   "Cooling System Operating" : Bool = PLC "68_Sys_Status_Data".CSW_IL_PRES_IN_RNG AT %DB1.DBX0.0, 1 s
   "Correct Phase Rotation" : Bool = PLC "10_DI_Data".MCCP_5PG1_OK AT %DB1.DBX0.0, 1 s
   "CSW Drain Valve Closed" : Bool = PLC "10_DI_Data".CV322_CLSD AT %DB1.DBX0.0, 1 s
   "CSW Drain Valve Control" : Bool = PLC "14_DQ_Data".CV321_322_CNTRL AT %DB1.DBX0.0, 1 s
   "CSW Drain Valve Open" : Bool = PLC "10_DI_Data".CV322_OPN AT %DB1.DBX0.0, 1 s
   "CSW Pump Control" : Bool = PLC "51_SLAVE_STATUS".P301_ENBLD AT %DB51.DBX14.3, 1 s
   "CSW Pump Enabled" : Bool = PLC "10 DI_DATA".P301_ENBLD AT %DB1.DBX0.0, 1 s
   "CSW Pump Tripped" : Bool = PLC "10 DI_DATA".P301_TRIPPED AT %DB1.DBX0.0, 1 s
   "CSW Valve Closed" : Bool = PLC "10_DI_Data".CV311_CLSD AT %DB1.DBW0, 1 s
   "CSW Valve Control" : Bool = PLC "14_DQ_Data".CV311_312_CNTRL AT %DB1.DBX0.0, 1 s
   "CSW Valve Open" : Bool = PLC "10_DI_Data".CV311_OPN AT %DB1.DBW0, 1 s
   "Current User" : WString[15] AT %DB1.DBX0.0
   "CV312 Present" : Bool = PLC "80_From_HMI".CV312_PRSNT AT %DB1.DBX0.0, 1 s
   "CV401 - IG Supply Valve Closed" : Bool = PLC "10_DI_Data".CV401_CLSD AT %DB1.DBX0.0, 1 s
   "CV401 - IG Supply Valve Control" : Bool = PLC "14_DQ_Data".CV401_CNTRL AT %DB1.DBX0.0, 1 s
   "CV401 - IG Supply Valve Opened" : Bool = PLC "10_DI_Data".CV401_OPN AT %DB1.DBX0.0, 1 s
   "CV403 - IG Vent Valve Position Feedback Scaled" : Real = PLC "12_AI_Data".CV403_SCALED AT %DB1.DBX0.0, 1 s
   "CV431 Present" : Bool = PLC "80_From_HMI".CV431_PRSNT AT %DB1.DBX0.0, 1 s
   "CV431/432 CB/BWTS Valve" : Bool = PLC "14_DQ_Data".CV431_432_CNTRL AT %DB1.DBX0.0, 1 s
   "CV432 Present" : Bool = PLC "80_From_HMI".CV432_PRSNT AT %DB1.DBX0.0, 1 s
   "Data To IGG PLC_Data_Fuel Oil System Proved" : Bool = PLC "68_Sys_Status_Data".FUEL_PRES_IN_RNG AT %DB1.DBX0.0, 1 s
   "Data To IGG PLC_Data_VSD Fault Flag" : Bool = PLC "10_DI_Data".E139_VSD_FLT AT %DB1.DBX0.0, 1 s
   "Data_From BC PLC_Data_IA Compressor Running" : Bool = PLC "68_Sys_Status_Data".IA_PRES_IN_RNG AT %DB1.DBX0.0, 1 s
   "Data_To_BC PLC_Data_Cooling Water System Proved" : Bool = PLC "10_DI_Data".CV311_OPN AT %DB1.DBX0.0, 1 s
   "db_time_sync_time_local_READ" : LDT = PLC db_time_sync_time_local_READ AT %M4.0, 1 s
   "db_time_sync_time_system_READ" : LDT = PLC db_time_sync_time_system_READ AT %M2.0, 1 s
   "DTB Valve Closed" : Bool = PLC "10_DI_Data".CV321_CLSD AT %DB1.DBX0.0, 1 s
   "DTB Valve Opened" : Bool = PLC "10_DI_Data".CV321_OPN AT %DB1.DBX0.0, 1 s
   "Evolving Setpoint_DB_LevelBetter" : Bool = PLC "Evolving Setpoint_DB".LevelBetter, 1 s
   "External Shutdown" : Bool = PLC "10 DI_DATA".ESD_OK AT %DB1.DBX0.0, 1 s
   "FDU Power Healthy" : Bool = PLC "10 DI_DATA".FD001_PWR_OK AT %DB1.DBX0.0, 1 s
   "FIT417_1S__ALM_ANALOG_DB_HIGH LEVEL VALUE (H)" : Real = PLC "FIT417_1S__ALM_ANALOG_DB"."HIGH LEVEL VALUE (H)" AT %DB2090.DBD30, 1 s
   "FIT417_1S__ALM_ANALOG_DB_LOW LEVEL VALUE (L)" : Real = PLC "FIT417_1S__ALM_ANALOG_DB"."LOW LEVEL VALUE (L)" AT %DB2090.DBD26, 1 s
   "FIT417_1S__ALM_ANALOG_DB_VERY HIGH LEVEL VALUE (HH)" : Real = PLC "FIT417_1S__ALM_ANALOG_DB"."VERY HIGH LEVEL VALUE (HH)" AT %DB2090.DBD34, 1 s
   "FIT417_1S__ALM_ANALOG_DB_VERY LOW LEVEL VALUE (LL)" : Real = PLC "FIT417_1S__ALM_ANALOG_DB"."VERY LOW LEVEL VALUE (LL)" AT %DB2090.DBD22, 1 s
   "FIT417_2S_ALM_ANALOG_DB_HIGH LEVEL VALUE (H)" : Real = PLC FIT417_2S_ALM_ANALOG_DB."HIGH LEVEL VALUE (H)" AT %DB2066.DBD30, 1 s
   "FIT417_2S_ALM_ANALOG_DB_LOW LEVEL VALUE (L)" : Real = PLC FIT417_2S_ALM_ANALOG_DB."LOW LEVEL VALUE (L)" AT %DB2066.DBD26, 1 s
   "FIT417_2S_ALM_ANALOG_DB_VERY HIGH LEVEL VALUE (HH)" : Real = PLC FIT417_2S_ALM_ANALOG_DB."VERY HIGH LEVEL VALUE (HH)" AT %DB2066.DBD34, 1 s
   "FIT417_2S_ALM_ANALOG_DB_VERY LOW LEVEL VALUE (LL)" : Real = PLC FIT417_2S_ALM_ANALOG_DB."VERY LOW LEVEL VALUE (LL)" AT %DB2066.DBD22, 1 s
   "FIT417_3S_ALM_ANALOG_DB_HIGH LEVEL VALUE (H)" : Real = PLC FIT417_3S_ALM_ANALOG_DB."HIGH LEVEL VALUE (H)" AT %DB2092.DBD30, 1 s
   "FIT417_3S_ALM_ANALOG_DB_LOW LEVEL VALUE (L)" : Real = PLC FIT417_3S_ALM_ANALOG_DB."LOW LEVEL VALUE (L)" AT %DB2092.DBD26, 1 s
   "FIT417_3S_ALM_ANALOG_DB_VERY HIGH LEVEL VALUE (HH)" : Real = PLC FIT417_3S_ALM_ANALOG_DB."VERY HIGH LEVEL VALUE (HH)" AT %DB2092.DBD34, 1 s
   "FIT417_3S_ALM_ANALOG_DB_VERY LOW LEVEL VALUE (LL)" : Real = PLC FIT417_3S_ALM_ANALOG_DB."VERY LOW LEVEL VALUE (LL)" AT %DB2092.DBD22, 1 s
   "FIT417_4S_ALM_ANALOG_DB_HIGH LEVEL VALUE (H)" : Real = PLC FIT417_4S_ALM_ANALOG_DB."HIGH LEVEL VALUE (H)" AT %DB2094.DBD30, 1 s
   "FIT417_4S_ALM_ANALOG_DB_LOW LEVEL VALUE (L)" : Real = PLC FIT417_4S_ALM_ANALOG_DB."LOW LEVEL VALUE (L)" AT %DB2094.DBD26, 1 s
   "FIT417_4S_ALM_ANALOG_DB_VERY HIGH LEVEL VALUE (HH)" : Real = PLC FIT417_4S_ALM_ANALOG_DB."VERY HIGH LEVEL VALUE (HH)" AT %DB2094.DBD34, 1 s
   "FIT417_4S_ALM_ANALOG_DB_VERY LOW LEVEL VALUE (LL)" : Real = PLC FIT417_4S_ALM_ANALOG_DB."VERY LOW LEVEL VALUE (LL)" AT %DB2094.DBD22, 1 s
   "FIT417_5S_ALM_ANALOG_DB_HIGH LEVEL VALUE (H)" : Real = PLC FIT417_5S_ALM_ANALOG_DB."HIGH LEVEL VALUE (H)" AT %DB2096.DBD30, 1 s
   "FIT417_5S_ALM_ANALOG_DB_LOW LEVEL VALUE (L)" : Real = PLC FIT417_5S_ALM_ANALOG_DB."LOW LEVEL VALUE (L)" AT %DB2096.DBD26, 1 s
   "FIT417_5S_ALM_ANALOG_DB_VERY HIGH LEVEL VALUE (HH)" : Real = PLC FIT417_5S_ALM_ANALOG_DB."VERY HIGH LEVEL VALUE (HH)" AT %DB2096.DBD34, 1 s
   "FIT417_5S_ALM_ANALOG_DB_VERY LOW LEVEL VALUE (LL)" : Real = PLC FIT417_5S_ALM_ANALOG_DB."VERY LOW LEVEL VALUE (LL)" AT %DB2096.DBD22, 1 s
   "FIT417_6S_ALM_ANALOG_DB_HIGH LEVEL VALUE (H)" : Real = PLC FIT417_6S_ALM_ANALOG_DB."HIGH LEVEL VALUE (H)" AT %DB2098.DBD30, 1 s
   "FIT417_6S_ALM_ANALOG_DB_LOW LEVEL VALUE (L)" : Real = PLC FIT417_6S_ALM_ANALOG_DB."LOW LEVEL VALUE (L)" AT %DB2098.DBD26, 1 s
   "FIT417_6S_ALM_ANALOG_DB_VERY HIGH LEVEL VALUE (HH)" : Real = PLC FIT417_6S_ALM_ANALOG_DB."VERY HIGH LEVEL VALUE (HH)" AT %DB2098.DBD34, 1 s
   "FIT417_6S_ALM_ANALOG_DB_VERY LOW LEVEL VALUE (LL)" : Real = PLC FIT417_6S_ALM_ANALOG_DB."VERY LOW LEVEL VALUE (LL)" AT %DB2098.DBD22, 1 s
   "FIT417_APT_ALM_ANALOG_DB_HIGH LEVEL VALUE (H)" : Real = PLC FIT417_APT_ALM_ANALOG_DB."HIGH LEVEL VALUE (H)" AT %DB2099.DBD30, 1 s
   "FIT417_APT_ALM_ANALOG_DB_LOW LEVEL VALUE (L)" : Real = PLC FIT417_APT_ALM_ANALOG_DB."LOW LEVEL VALUE (L)" AT %DB2099.DBD26, 1 s
   "FIT417_APT_ALM_ANALOG_DB_VERY HIGH LEVEL VALUE (HH)" : Real = PLC FIT417_APT_ALM_ANALOG_DB."VERY HIGH LEVEL VALUE (HH)" AT %DB2099.DBD34, 1 s
   "FIT417_APT_ALM_ANALOG_DB_VERY LOW LEVEL VALUE (LL)" : Real = PLC FIT417_APT_ALM_ANALOG_DB."VERY LOW LEVEL VALUE (LL)" AT %DB2099.DBD22, 1 s
   "FIT418_1P__ALM_ANALOG_DB_HIGH LEVEL VALUE (H)" : Real = PLC "FIT418_1P__ALM_ANALOG_DB"."HIGH LEVEL VALUE (H)" AT %DB2089.DBD30, 1 s
   "FIT418_1P__ALM_ANALOG_DB_LOW LEVEL VALUE (L)" : Real = PLC "FIT418_1P__ALM_ANALOG_DB"."LOW LEVEL VALUE (L)" AT %DB2089.DBD26, 1 s
   "FIT418_1P__ALM_ANALOG_DB_VERY HIGH LEVEL VALUE (HH)" : Real = PLC "FIT418_1P__ALM_ANALOG_DB"."VERY HIGH LEVEL VALUE (HH)" AT %DB2089.DBD34, 1 s
   "FIT418_1P__ALM_ANALOG_DB_VERY LOW LEVEL VALUE (LL)" : Real = PLC "FIT418_1P__ALM_ANALOG_DB"."VERY LOW LEVEL VALUE (LL)" AT %DB2089.DBD22, 1 s
   "FIT418_2P_ALM_ANALOG_DB_ALARM L" : Bool = PLC FIT418_2P_ALM_ANALOG_DB."ALARM L" AT %DB2064.DBX48.2, 1 s
   "FIT418_2P_ALM_ANALOG_DB_HIGH LEVEL VALUE (H)" : Real = PLC FIT418_2P_ALM_ANALOG_DB."HIGH LEVEL VALUE (H)" AT %DB2064.DBD30, 1 s
   "FIT418_2P_ALM_ANALOG_DB_LOW LEVEL VALUE (L)" : Real = PLC FIT418_2P_ALM_ANALOG_DB."LOW LEVEL VALUE (L)" AT %DB2064.DBD26, 1 s
   "FIT418_2P_ALM_ANALOG_DB_VERY HIGH LEVEL VALUE (HH)" : Real = PLC FIT418_2P_ALM_ANALOG_DB."VERY HIGH LEVEL VALUE (HH)" AT %DB2064.DBD34, 1 s
   "FIT418_2P_ALM_ANALOG_DB_VERY LOW LEVEL VALUE (LL)" : Real = PLC FIT418_2P_ALM_ANALOG_DB."VERY LOW LEVEL VALUE (LL)" AT %DB2064.DBD22, 1 s
   "FIT418_3P__ALM_ANALOG_DB_HIGH LEVEL VALUE (H)" : Real = PLC "FIT418_3P__ALM_ANALOG_DB"."HIGH LEVEL VALUE (H)" AT %DB2091.DBD30, 1 s
   "FIT418_3P__ALM_ANALOG_DB_LOW LEVEL VALUE (L)" : Real = PLC "FIT418_3P__ALM_ANALOG_DB"."LOW LEVEL VALUE (L)" AT %DB2091.DBD26, 1 s
   "FIT418_3P__ALM_ANALOG_DB_VERY HIGH LEVEL VALUE (HH)" : Real = PLC "FIT418_3P__ALM_ANALOG_DB"."VERY HIGH LEVEL VALUE (HH)" AT %DB2091.DBD34, 1 s
   "FIT418_3P__ALM_ANALOG_DB_VERY LOW LEVEL VALUE (LL)" : Real = PLC "FIT418_3P__ALM_ANALOG_DB"."VERY LOW LEVEL VALUE (LL)" AT %DB2091.DBD22, 1 s
   "FIT418_4P__ALM_ANALOG_DB_HIGH LEVEL VALUE (H)" : Real = PLC "FIT418_4P__ALM_ANALOG_DB"."HIGH LEVEL VALUE (H)" AT %DB2093.DBD30, 1 s
   "FIT418_4P__ALM_ANALOG_DB_LOW LEVEL VALUE (L)" : Real = PLC "FIT418_4P__ALM_ANALOG_DB"."LOW LEVEL VALUE (L)" AT %DB2093.DBD26, 1 s
   "FIT418_4P__ALM_ANALOG_DB_VERY HIGH LEVEL VALUE (HH)" : Real = PLC "FIT418_4P__ALM_ANALOG_DB"."VERY HIGH LEVEL VALUE (HH)" AT %DB2093.DBD34, 1 s
   "FIT418_4P__ALM_ANALOG_DB_VERY LOW LEVEL VALUE (LL)" : Real = PLC "FIT418_4P__ALM_ANALOG_DB"."VERY LOW LEVEL VALUE (LL)" AT %DB2093.DBD22, 1 s
   "FIT418_5P__ALM_ANALOG_DB_HIGH LEVEL VALUE (H)" : Real = PLC "FIT418_5P__ALM_ANALOG_DB"."HIGH LEVEL VALUE (H)" AT %DB2095.DBD30, 1 s
   "FIT418_5P__ALM_ANALOG_DB_LOW LEVEL VALUE (L)" : Real = PLC "FIT418_5P__ALM_ANALOG_DB"."LOW LEVEL VALUE (L)" AT %DB2095.DBD26, 1 s
   "FIT418_5P__ALM_ANALOG_DB_VERY HIGH LEVEL VALUE (HH)" : Real = PLC "FIT418_5P__ALM_ANALOG_DB"."VERY HIGH LEVEL VALUE (HH)" AT %DB2095.DBD34, 1 s
   "FIT418_5P__ALM_ANALOG_DB_VERY LOW LEVEL VALUE (LL)" : Real = PLC "FIT418_5P__ALM_ANALOG_DB"."VERY LOW LEVEL VALUE (LL)" AT %DB2095.DBD22, 1 s
   "FIT418_6P__ALM_ANALOG_DB_HIGH LEVEL VALUE (H)" : Real = PLC "FIT418_6P__ALM_ANALOG_DB"."HIGH LEVEL VALUE (H)" AT %DB2097.DBD30, 1 s
   "FIT418_6P__ALM_ANALOG_DB_LOW LEVEL VALUE (L)" : Real = PLC "FIT418_6P__ALM_ANALOG_DB"."LOW LEVEL VALUE (L)" AT %DB2097.DBD26, 1 s
   "FIT418_6P__ALM_ANALOG_DB_VERY HIGH LEVEL VALUE (HH)" : Real = PLC "FIT418_6P__ALM_ANALOG_DB"."VERY HIGH LEVEL VALUE (HH)" AT %DB2097.DBD34, 1 s
   "FIT418_6P__ALM_ANALOG_DB_VERY LOW LEVEL VALUE (LL)" : Real = PLC "FIT418_6P__ALM_ANALOG_DB"."VERY LOW LEVEL VALUE (LL)" AT %DB2097.DBD22, 1 s
   "FIT418_FPT__ALM_ANALOG_DB_HIGH LEVEL VALUE (H)" : Real = PLC "FIT418_FPT__ALM_ANALOG_DB"."HIGH LEVEL VALUE (H)" AT %DB2088.DBD30, 1 s
   "FIT418_FPT__ALM_ANALOG_DB_LOW LEVEL VALUE (L)" : Real = PLC "FIT418_FPT__ALM_ANALOG_DB"."LOW LEVEL VALUE (L)" AT %DB2088.DBD26, 1 s
   "FIT418_FPT__ALM_ANALOG_DB_VERY HIGH LEVEL VALUE (HH)" : Real = PLC "FIT418_FPT__ALM_ANALOG_DB"."VERY HIGH LEVEL VALUE (HH)" AT %DB2088.DBD34, 1 s
   "FIT418_FPT__ALM_ANALOG_DB_VERY LOW LEVEL VALUE (LL)" : Real = PLC "FIT418_FPT__ALM_ANALOG_DB"."VERY LOW LEVEL VALUE (LL)" AT %DB2088.DBD22, 1 s
   "FIT419_ALM_ANALOG_DB_HIGH LEVEL VALUE (H)" : Real = PLC FIT419_ALM_ANALOG_DB."HIGH LEVEL VALUE (H)" AT %DB2067.DBD30, 1 s
   "FIT419_ALM_ANALOG_DB_LOW LEVEL VALUE (L)" : Real = PLC FIT419_ALM_ANALOG_DB."LOW LEVEL VALUE (L)" AT %DB2067.DBD26, 1 s
   "FIT419_ALM_ANALOG_DB_VERY HIGH LEVEL VALUE (HH)" : Real = PLC FIT419_ALM_ANALOG_DB."VERY HIGH LEVEL VALUE (HH)" AT %DB2067.DBD34, 1 s
   "FIT419_ALM_ANALOG_DB_VERY LOW LEVEL VALUE (LL)" : Real = PLC FIT419_ALM_ANALOG_DB."VERY LOW LEVEL VALUE (LL)" AT %DB2067.DBD22, 1 s
   "FIT420_1P_ALM_ANALOG_DB_HIGH LEVEL VALUE (H)" : Real = PLC FIT420_1P_ALM_ANALOG_DB."HIGH LEVEL VALUE (H)" AT %DB2202.DBD30, 1 s
   "FIT420_1P_ALM_ANALOG_DB_LOW LEVEL VALUE (L)" : Real = PLC FIT420_1P_ALM_ANALOG_DB."LOW LEVEL VALUE (L)" AT %DB2202.DBD26, 1 s
   "FIT420_1P_ALM_ANALOG_DB_VERY HIGH LEVEL VALUE (HH)" : Real = PLC FIT420_1P_ALM_ANALOG_DB."VERY HIGH LEVEL VALUE (HH)" AT %DB2202.DBD34, 1 s
   "FIT420_1P_ALM_ANALOG_DB_VERY LOW LEVEL VALUE (LL)" : Real = PLC FIT420_1P_ALM_ANALOG_DB."VERY LOW LEVEL VALUE (LL)" AT %DB2202.DBD22, 1 s
   "FIT420_1S_ALM_ANALOG_DB_HIGH LEVEL VALUE (H)" : Real = PLC FIT420_1S_ALM_ANALOG_DB."HIGH LEVEL VALUE (H)" AT %DB2203.DBD30, 1 s
   "FIT420_1S_ALM_ANALOG_DB_LOW LEVEL VALUE (L)" : Real = PLC FIT420_1S_ALM_ANALOG_DB."LOW LEVEL VALUE (L)" AT %DB2203.DBD26, 1 s
   "FIT420_1S_ALM_ANALOG_DB_VERY HIGH LEVEL VALUE (HH)" : Real = PLC FIT420_1S_ALM_ANALOG_DB."VERY HIGH LEVEL VALUE (HH)" AT %DB2203.DBD34, 1 s
   "FIT420_1S_ALM_ANALOG_DB_VERY LOW LEVEL VALUE (LL)" : Real = PLC FIT420_1S_ALM_ANALOG_DB."VERY LOW LEVEL VALUE (LL)" AT %DB2203.DBD22, 1 s
   "FIT420_3P_ALM_ANALOG_DB_HIGH LEVEL VALUE (H)" : Real = PLC FIT420_3P_ALM_ANALOG_DB."HIGH LEVEL VALUE (H)" AT %DB2204.DBD30, 1 s
   "FIT420_3P_ALM_ANALOG_DB_LOW LEVEL VALUE (L)" : Real = PLC FIT420_3P_ALM_ANALOG_DB."LOW LEVEL VALUE (L)" AT %DB2204.DBD26, 1 s
   "FIT420_3P_ALM_ANALOG_DB_VERY HIGH LEVEL VALUE (HH)" : Real = PLC FIT420_3P_ALM_ANALOG_DB."VERY HIGH LEVEL VALUE (HH)" AT %DB2204.DBD34, 1 s
   "FIT420_3P_ALM_ANALOG_DB_VERY LOW LEVEL VALUE (LL)" : Real = PLC FIT420_3P_ALM_ANALOG_DB."VERY LOW LEVEL VALUE (LL)" AT %DB2204.DBD22, 1 s
   "FIT420_3S_ALM_ANALOG_DB_HIGH LEVEL VALUE (H)" : Real = PLC FIT420_3S_ALM_ANALOG_DB."HIGH LEVEL VALUE (H)" AT %DB2205.DBD30, 1 s
   "FIT420_3S_ALM_ANALOG_DB_LOW LEVEL VALUE (L)" : Real = PLC FIT420_3S_ALM_ANALOG_DB."LOW LEVEL VALUE (L)" AT %DB2205.DBD26, 1 s
   "FIT420_3S_ALM_ANALOG_DB_VERY HIGH LEVEL VALUE (HH)" : Real = PLC FIT420_3S_ALM_ANALOG_DB."VERY HIGH LEVEL VALUE (HH)" AT %DB2205.DBD34, 1 s
   "FIT420_3S_ALM_ANALOG_DB_VERY LOW LEVEL VALUE (LL)" : Real = PLC FIT420_3S_ALM_ANALOG_DB."VERY LOW LEVEL VALUE (LL)" AT %DB2205.DBD22, 1 s
   "FIT420_4P_ALM_ANALOG_DB_HIGH LEVEL VALUE (H)" : Real = PLC FIT420_4P_ALM_ANALOG_DB."HIGH LEVEL VALUE (H)" AT %DB2206.DBD30, 1 s
   "FIT420_4P_ALM_ANALOG_DB_LOW LEVEL VALUE (L)" : Real = PLC FIT420_4P_ALM_ANALOG_DB."LOW LEVEL VALUE (L)" AT %DB2206.DBD26, 1 s
   "FIT420_4P_ALM_ANALOG_DB_VERY HIGH LEVEL VALUE (HH)" : Real = PLC FIT420_4P_ALM_ANALOG_DB."VERY HIGH LEVEL VALUE (HH)" AT %DB2206.DBD34, 1 s
   "FIT420_4P_ALM_ANALOG_DB_VERY LOW LEVEL VALUE (LL)" : Real = PLC FIT420_4P_ALM_ANALOG_DB."VERY LOW LEVEL VALUE (LL)" AT %DB2206.DBD22, 1 s
   "FIT420_4S_ALM_ANALOG_DB_HIGH LEVEL VALUE (H)" : Real = PLC FIT420_4S_ALM_ANALOG_DB."HIGH LEVEL VALUE (H)" AT %DB2207.DBD30, 1 s
   "FIT420_4S_ALM_ANALOG_DB_LOW LEVEL VALUE (L)" : Real = PLC FIT420_4S_ALM_ANALOG_DB."LOW LEVEL VALUE (L)" AT %DB2207.DBD26, 1 s
   "FIT420_4S_ALM_ANALOG_DB_VERY HIGH LEVEL VALUE (HH)" : Real = PLC FIT420_4S_ALM_ANALOG_DB."VERY HIGH LEVEL VALUE (HH)" AT %DB2207.DBD34, 1 s
   "FIT420_4S_ALM_ANALOG_DB_VERY LOW LEVEL VALUE (LL)" : Real = PLC FIT420_4S_ALM_ANALOG_DB."VERY LOW LEVEL VALUE (LL)" AT %DB2207.DBD22, 1 s
   "FIT420_5P_ALM_ANALOG_DB_HIGH LEVEL VALUE (H)" : Real = PLC FIT420_5P_ALM_ANALOG_DB."HIGH LEVEL VALUE (H)" AT %DB2208.DBD30, 1 s
   "FIT420_5P_ALM_ANALOG_DB_LOW LEVEL VALUE (L)" : Real = PLC FIT420_5P_ALM_ANALOG_DB."LOW LEVEL VALUE (L)" AT %DB2208.DBD26, 1 s
   "FIT420_5P_ALM_ANALOG_DB_VERY HIGH LEVEL VALUE (HH)" : Real = PLC FIT420_5P_ALM_ANALOG_DB."VERY HIGH LEVEL VALUE (HH)" AT %DB2208.DBD34, 1 s
   "FIT420_5P_ALM_ANALOG_DB_VERY LOW LEVEL VALUE (LL)" : Real = PLC FIT420_5P_ALM_ANALOG_DB."VERY LOW LEVEL VALUE (LL)" AT %DB2208.DBD22, 1 s
   "FIT420_5S_ALM_ANALOG_DB_HIGH LEVEL VALUE (H)" : Real = PLC FIT420_5S_ALM_ANALOG_DB."HIGH LEVEL VALUE (H)" AT %DB2209.DBD30, 1 s
   "FIT420_5S_ALM_ANALOG_DB_LOW LEVEL VALUE (L)" : Real = PLC FIT420_5S_ALM_ANALOG_DB."LOW LEVEL VALUE (L)" AT %DB2209.DBD26, 1 s
   "FIT420_5S_ALM_ANALOG_DB_VERY HIGH LEVEL VALUE (HH)" : Real = PLC FIT420_5S_ALM_ANALOG_DB."VERY HIGH LEVEL VALUE (HH)" AT %DB2209.DBD34, 1 s
   "FIT420_5S_ALM_ANALOG_DB_VERY LOW LEVEL VALUE (LL)" : Real = PLC FIT420_5S_ALM_ANALOG_DB."VERY LOW LEVEL VALUE (LL)" AT %DB2209.DBD22, 1 s
   "FIT420_6P_ALM_ANALOG_DB_HIGH LEVEL VALUE (H)" : Real = PLC FIT420_6P_ALM_ANALOG_DB."HIGH LEVEL VALUE (H)" AT %DB2210.DBD30, 1 s
   "FIT420_6P_ALM_ANALOG_DB_LOW LEVEL VALUE (L)" : Real = PLC FIT420_6P_ALM_ANALOG_DB."LOW LEVEL VALUE (L)" AT %DB2210.DBD26, 1 s
   "FIT420_6P_ALM_ANALOG_DB_VERY HIGH LEVEL VALUE (HH)" : Real = PLC FIT420_6P_ALM_ANALOG_DB."VERY HIGH LEVEL VALUE (HH)" AT %DB2210.DBD34, 1 s
   "FIT420_6P_ALM_ANALOG_DB_VERY LOW LEVEL VALUE (LL)" : Real = PLC FIT420_6P_ALM_ANALOG_DB."VERY LOW LEVEL VALUE (LL)" AT %DB2210.DBD22, 1 s
   "FIT420_6S_ALM_ANALOG_DB_HIGH LEVEL VALUE (H)" : Real = PLC FIT420_6S_ALM_ANALOG_DB."HIGH LEVEL VALUE (H)" AT %DB2211.DBD30, 1 s
   "FIT420_6S_ALM_ANALOG_DB_LOW LEVEL VALUE (L)" : Real = PLC FIT420_6S_ALM_ANALOG_DB."LOW LEVEL VALUE (L)" AT %DB2211.DBD26, 1 s
   "FIT420_6S_ALM_ANALOG_DB_VERY HIGH LEVEL VALUE (HH)" : Real = PLC FIT420_6S_ALM_ANALOG_DB."VERY HIGH LEVEL VALUE (HH)" AT %DB2211.DBD34, 1 s
   "FIT420_6S_ALM_ANALOG_DB_VERY LOW LEVEL VALUE (LL)" : Real = PLC FIT420_6S_ALM_ANALOG_DB."VERY LOW LEVEL VALUE (LL)" AT %DB2211.DBD22, 1 s
   "FIT420_APT_ALM_ANALOG_DB_HIGH LEVEL VALUE (H)" : Real = PLC FIT420_APT_ALM_ANALOG_DB."HIGH LEVEL VALUE (H)" AT %DB2212.DBD30, 1 s
   "FIT420_APT_ALM_ANALOG_DB_LOW LEVEL VALUE (L)" : Real = PLC FIT420_APT_ALM_ANALOG_DB."LOW LEVEL VALUE (L)" AT %DB2212.DBD26, 1 s
   "FIT420_APT_ALM_ANALOG_DB_VERY HIGH LEVEL VALUE (HH)" : Real = PLC FIT420_APT_ALM_ANALOG_DB."VERY HIGH LEVEL VALUE (HH)" AT %DB2212.DBD34, 1 s
   "FIT420_APT_ALM_ANALOG_DB_VERY LOW LEVEL VALUE (LL)" : Real = PLC FIT420_APT_ALM_ANALOG_DB."VERY LOW LEVEL VALUE (LL)" AT %DB2212.DBD22, 1 s
   "FIT420_FPT_ALM_ANALOG_DB_HIGH LEVEL VALUE (H)" : Real = PLC FIT420_FPT_ALM_ANALOG_DB."HIGH LEVEL VALUE (H)" AT %DB2201.DBD30, 1 s
   "FIT420_FPT_ALM_ANALOG_DB_LOW LEVEL VALUE (L)" : Real = PLC FIT420_FPT_ALM_ANALOG_DB."LOW LEVEL VALUE (L)" AT %DB2201.DBD26, 1 s
   "FIT420_FPT_ALM_ANALOG_DB_VERY HIGH LEVEL VALUE (HH)" : Real = PLC FIT420_FPT_ALM_ANALOG_DB."VERY HIGH LEVEL VALUE (HH)" AT %DB2201.DBD34, 1 s
   "FIT420_FPT_ALM_ANALOG_DB_VERY LOW LEVEL VALUE (LL)" : Real = PLC FIT420_FPT_ALM_ANALOG_DB."VERY LOW LEVEL VALUE (LL)" AT %DB2201.DBD22, 1 s
   "FIT420PORT_ALM_ANALOG_DB_HIGH LEVEL VALUE (H)" : Real = PLC FIT420PORT_ALM_ANALOG_DB."HIGH LEVEL VALUE (H)" AT %DB2065.DBD30, 1 s
   "FIT420PORT_ALM_ANALOG_DB_LOW LEVEL VALUE (L)" : Real = PLC FIT420PORT_ALM_ANALOG_DB."LOW LEVEL VALUE (L)" AT %DB2065.DBD26, 1 s
   "FIT420PORT_ALM_ANALOG_DB_VERY HIGH LEVEL VALUE (HH)" : Real = PLC FIT420PORT_ALM_ANALOG_DB."VERY HIGH LEVEL VALUE (HH)" AT %DB2065.DBD34, 1 s
   "FIT420PORT_ALM_ANALOG_DB_VERY LOW LEVEL VALUE (LL)" : Real = PLC FIT420PORT_ALM_ANALOG_DB."VERY LOW LEVEL VALUE (LL)" AT %DB2065.DBD22, 1 s
   "Flame" : Bool = PLC "103_Main_Burner_DB".DN_OK AT %DB1.DBX0.0, 1 s
   "Flame Signal OK" : Bool = PLC "10 DI_DATA".FD001_OK AT %DB1.DBX0.0, 1 s
   "Flame Signal Scaled" : Real = PLC "12_AI_Data".FD001FlameSignalIn AT %DB1.DBX0.0, 100 ms
   "Flue gas Scrubber Valve Closed" : Bool = PLC "10_DI_Data".CV312_CLSD AT %DB1.DBX0.0, 1 s
   "Flue Gas Scrubber Valve Opened" : Bool = PLC "10_DI_Data".CV312_OPN AT %DB1.DBX0.0, 1 s
   "FP1 Running" : Bool = PLC "10_DI_Data".E500A_ENBLD AT %DB1.DBX0.0, 1 s
   "FP2 Running" : Bool = PLC "10_DI_Data".E500B_ENBLD AT %DB1.DBX0.0, 1 s
   "FPT BWT Level High High Switch" : Bool = PLC "FPT BWT Level High High Switch" AT %I9.0, 1 s
   "FPT GTT Isolation Valve Feedback - Closed" : Bool = PLC "FPT GTT Isolation Valve Feedback - Closed" AT %I0.1, 1 s
   "FPT GTT Isolation Valve Feedback - Opened" : Bool = PLC "FPT GTT Isolation Valve Feedback - Opened" AT %I0.0, 1 s
   "FPT Tank Vent Valve 1 Feedback - Closed" : Bool = PLC "FPT Tank Vent Valve 1 Feedback - Closed" AT %I0.3, 1 s
   "FPT Tank Vent Valve 1 Feedback - Opened" : Bool = PLC "FPT Tank Vent Valve 1 Feedback - Opened" AT %I0.2, 1 s
   "FPT Tank Vent Valve 2 Feedback - Closed" : Bool = PLC "FPT Tank Vent Valve 2 Feedback - Closed" AT %I0.5, 1 s
   "FPT Tank Vent Valve 2 Feedback - Opened" : Bool = PLC "FPT Tank Vent Valve 2 Feedback - Opened" AT %I0.4, 1 s
   "Fresh Water Bulk Tank Level (LIT305) Scaled" : Real = PLC "12_AI_Data".LIT305_SCALED AT %DB1.DBX0.0, 1 s
   "Fresh Water Pump Control" : Bool = PLC "14_DQ_Data".P305ControlOut AT %DB1.DBX0.0, 1 s
   "Fresh Water Pump Enabled" : Bool = PLC "10 DI_DATA".P305_ENBLD AT %DB1.DBX0.0, 1 s
   "Fresh Water Pump Enabled(1)" : Bool = PLC "10 DI_DATA".P305_ENBLD AT %DB1.DBX0.0, 1 s
   "Fresh Water Pump Run Minutes" : Int = PLC "P305_Functioning Hours_IDB".Minutes, 1 s
   "Fresh Water Pump Run Seconds" : Int = PLC "P305_Functioning Hours_IDB".Seconds, 1 s
   "Fresh Water Pump Service Due" : Bool = PLC "P305_Functioning Hours_IDB"."Service Time bit", 1 s
   "Fresh Water Pump Total Run Hours" : Int = PLC "P305_Functioning Hours_IDB"."Hours Total", 1 s
   "Fresh Water Pump Tripped" : Bool = PLC "10 DI_DATA".P305_TRIPPED AT %DB1.DBX0.0, 1 s
   "Fresh Water Pump Tripped Alarm" : Bool = PLC "10 DI_DATA".P305_TRIPPED AT %DB1.DBX0.0, 1 s
   "Fuel Pressure Setting" : Real = PLC "84_Setpoints".PIT205_Target AT %DB1.DBX0.0, 1 s
   "Fuel Pump 1 Animation" : Int = PLC "82_To_HMI"."Fuel Pump 1 Animation", 1 s
   "Fuel Pump 1 Control" : Bool = PLC "14_DQ_Data".E500A_CNTRL AT %DB1.DBX0.0, 1 s
   "Fuel Pump 1 Enabled" : Bool = PLC "10_DI_Data".E500A_ENBLD AT %DB1.DBX0.0, 1 s
   "Fuel Pump 1 Tripped" : Bool = PLC "10_DI_Data".E500A_TRIPPED AT %DB1.DBX0.0, 1 s
   "Fuel Pump 2 Animation" : Int = PLC "82_To_HMI"."Fuel Pump 2 Animation", 1 s
   "Fuel Pump 2 Control" : Bool = PLC "14_DQ_Data".E500B_CNTRL AT %DB1.DBX0.0, 1 s
   "Fuel Pump 2 Enabled" : Bool = PLC "10_DI_Data".E500B_ENBLD AT %DB1.DBX0.0, 1 s
   "Fuel Pump 2 Fault" : Bool = PLC "10_DI_Data".E500B_TRIPPED AT %DB1.DBX0.0, 1 s
   "Fuel Pump 2 Tripped" : Bool = PLC "10_DI_Data".E500B_TRIPPED AT %DB1.DBX0.0, 1 s
   "Fuel Valve Manual Regulator" : Int, internal
   "FW Pump Animation" : Int, internal
   "HMI Ballast Water Treatment" : Bool = PLC "80_From_HMI".BWT_BYPASS AT %DB1.DBX0.0, 1 s
   "HMI Cargo Blanketing" : Bool = PLC "80_From_HMI".CRG_BLNK_MODE AT %DB1.DBX0.0, 1 s
   "HMI Data_Atmospheric Oxygen 1 Low" : Real = PLC "84_Setpoints".AT_O2_1_Low AT %DB1.DBD0, 1 s
   "HMI Data_Atmospheric Oxygen 1 Low Low" : Real = PLC "84_Setpoints".AT_O2_1_LowLow AT %DB1.DBD0, 1 s
   "HMI Data_Atmospheric Oxygen 2 Low" : Real = PLC "84_Setpoints".AT_O2_2_Low AT %DB1.DBD0, 1 s
   "HMI Data_Atmospheric Oxygen 2 Low Low" : Real = PLC "84_Setpoints".AT_O2_2_LowLow AT %DB1.DBD0, 1 s
   "HMI Data_Atomising Air Preassure High High" : Real = PLC "84_Setpoints".PIT113_HighHigh AT %DB1.DBD0, 1 s
   "HMI Data_Atomising Air Preassure Low Low SP" : Real = PLC "84_Setpoints".PIT113_LowLow AT %DB1.DBD0, 1 s
   "HMI Data_Atomising Air Pressure High" : Real = PLC "84_Setpoints".PIT113_High AT %DB1.DBD0, 1 s
   "HMI Data_Atomising Air Pressure Low SP" : Real = PLC "84_Setpoints".PIT113_Low AT %DB1.DBD0, 1 s
   "HMI Data_Atomising Air Reg Pressure Setpoint" : Real = PLC "84_Setpoints".PIT113_Pilot_Target AT %DB1.DBX0.0, 1 s
   "HMI Data_Blower Service Time" : Int = PLC "82_To_HMI"."CA Blower Service Time Hours", 1 s
   "HMI Data_CA Blower Pressure(PIT102) High" : Real = PLC "84_Setpoints".PIT102_Main_High AT %DB1.DBD0, 1 s
   "HMI Data_CA Blower Pressure(PIT102) High High" : Real = PLC "84_Setpoints".PIT102_Main_HighHigh AT %DB1.DBD0, 1 s
   "HMI Data_CA Blower Pressure(PIT102) High High_Post" : Real = PLC "84_Setpoints".PIT102_Post_HighHigh AT %DB1.DBD0, 1 s
   "HMI Data_CA Blower Pressure(PIT102) High High_Pre-Ignition" : Real = PLC "84_Setpoints".PIT102_Pilot_HighHigh AT %DB1.DBD0, 1 s
   "HMI Data_CA Blower Pressure(PIT102) High_Post" : Real = PLC "84_Setpoints".PIT102_Post_High AT %DB1.DBD0, 1 s
   "HMI Data_CA Blower Pressure(PIT102) High_Pre-Ignition" : Real = PLC "84_Setpoints".PIT102_Pilot_High AT %DB1.DBD0, 1 s
   "HMI Data_CA Blower Pressure(PIT102) Low" : Real = PLC "84_Setpoints".PIT102_Main_Low AT %DB1.DBD0, 1 s
   "HMI Data_CA Blower Pressure(PIT102) Low Low" : Real = PLC "84_Setpoints".PIT102_Main_LowLow AT %DB1.DBD0, 1 s
   "HMI Data_CA Blower Pressure(PIT102) Low Low_Post" : Real = PLC "84_Setpoints".PIT102_Post_LowLow AT %DB1.DBD0, 1 s
   "HMI Data_CA Blower Pressure(PIT102) Low Low_Pre-Ignition" : Real = PLC "84_Setpoints".PIT102_Pilot_LowLow AT %DB1.DBX0.0, 1 s
   "HMI Data_CA Blower Pressure(PIT102) Low_Post" : Real = PLC "84_Setpoints".PIT102_Post_Low AT %DB1.DBD0, 1 s
   "HMI Data_CA Blower Pressure(PIT102) Low_Pre-Ignition" : Real = PLC "84_Setpoints".PIT102_Pilot_Low AT %DB1.DBX0.0, 1 s
   "HMI Data_CA Start Up Press SP" : Real = PLC "84_Setpoints".PIT402_Pilot_Target AT %DB1.DBD0, 1 s
   "HMI Data_Cooling System Overrun" : Time = PLC "80_From_HMI"."Cooling System Overrun", 1 s
   "HMI Data_CSW Inlet Temp High" : Real = PLC "84_Setpoints".TIT319_High AT %DB1.DBD0, 1 s
   "HMI Data_CSW Inlet Temp High High" : Real = PLC "84_Setpoints".TIT319_HighHigh AT %DB1.DBD0, 1 s
   "HMI Data_CSW Oulet Temp High" : Real = PLC "84_Setpoints".TIT360_High AT %DB1.DBD0, 1 s
   "HMI Data_CSW Oulet Temp High High" : Real = PLC "84_Setpoints".TIT360_HighHigh AT %DB1.DBD0, 1 s
   "HMI Data_E600 BWTS Target" : Real = PLC "84_Setpoints".E600_BWT_Target AT %DB1.DBD0, 1 s
   "HMI Data_E600 CB Target" : Real = PLC "84_Setpoints".E600_CB_Target AT %DB1.DBD0, 1 s
   "HMI Data_FD001 Target" : Real = PLC "84_Setpoints".FD001_Min AT %DB1.DBD0, 1 s
   "HMI Data_Flame Signal Low" : Real = PLC "84_Setpoints".FD001_Low AT %DB1.DBD0, 1 s
   "HMI Data_Flame Signal Low Low" : Real = PLC "84_Setpoints".FD001_LowLow AT %DB1.DBD0, 1 s
   "HMI Data_Fresh Water Service Time" : Int = PLC "82_To_HMI"."P305 FW Pump Service Time Hours", 1 s
   "HMI Data_Fuel Pump Service Time" : LTime = PLC "80_From_HMI".MAX_E500_RT AT %DB1.DBX0.0, 1 s
   "HMI Data_HMI Blower Speed" : Real = PLC "80_From_HMI".E139_SET_SPEED AT %DB1.DBX0.0, 1 s
   "HMI Data_I&A Compressor Service Time" : Int = PLC "82_To_HMI"."I&A Compressor Service Time Hours", 1 s
   "HMI Data_IG O2 High BWTS" : Real = PLC "84_Setpoints".E600_BWT_High AT %DB1.DBD0, 1 s
   "HMI Data_IG O2 High CB" : Real = PLC "84_Setpoints".E600_CB_High AT %DB1.DBD0, 1 s
   "HMI Data_IG O2 High High BWTS" : Real = PLC "84_Setpoints".E600_BWT_HighHigh AT %DB1.DBD0, 1 s
   "HMI Data_IG O2 High High CB" : Real = PLC "84_Setpoints".E600_CB_HighHigh AT %DB1.DBD0, 1 s
   "HMI Data_IG O2 Low BWTS" : Real = PLC "84_Setpoints".E600_BWT_Low AT %DB1.DBD0, 1 s
   "HMI Data_IG O2 Low CB" : Real = PLC "84_Setpoints".E600_CB_Low AT %DB1.DBD0, 1 s
   "HMI Data_IG O2 Low Low BWTS" : Real = PLC "84_Setpoints".E600_BWT_LowLow AT %DB1.DBD0, 1 s
   "HMI Data_IG O2 Low Low CB" : Real = PLC "84_Setpoints".E600_CB_LowLow AT %DB1.DBD0, 1 s
   "HMI Data_IGG Inlet Fuel Pressure High" : Real = PLC "84_Setpoints".PIT204_High, 1 s
   "HMI Data_IGG Inlet Fuel Pressure High High" : Real = PLC "84_Setpoints".PIT204_HighHigh, 1 s
   "HMI Data_IGG Inlet Fuel Pressure Low Low SP" : Real = PLC "84_Setpoints".PIT204_LowLow, 1 s
   "HMI Data_IGG Inlet Fuel Pressure Low SP" : Real = PLC "84_Setpoints".PIT204_Low, 1 s
   "HMI Data_IGG Inlet Fuel Temperature High" : Real = PLC "84_Setpoints".TIT202_High AT %DB1.DBD0, 1 s
   "HMI Data_IGG Inlet Fuel Temperature High High" : Real = PLC "84_Setpoints".TIT202_HighHigh AT %DB1.DBD0, 1 s
   "HMI Data_IGG Inlet Fuel Temperature Low" : Real = PLC "84_Setpoints".TIT202_Low AT %DB1.DBD0, 1 s
   "HMI Data_IGG Inlet Fuel Temperature Low Low" : Real = PLC "84_Setpoints".TIT202_LowLow AT %DB1.DBD0, 1 s
   "HMI Data_IGG Pressure Setpoint" : Real = PLC "84_Setpoints".PIT402_Main_Target AT %DB1.DBX0.0, 1 s
   "HMI Data_Inert Gas Pressure (PIT402) High" : Real = PLC "84_Setpoints".PIT402_Main_High AT %DB1.DBD0, 1 s
   "HMI Data_Inert Gas Pressure (PIT402) High High" : Real = PLC "84_Setpoints".PIT402_Main_HighHigh AT %DB1.DBD0, 1 s
   "HMI Data_Inert Gas Pressure (PIT402) High High_Post" : Real = PLC "84_Setpoints".PIT402_Post_HighHigh AT %DB1.DBD0, 1 s
   "HMI Data_Inert Gas Pressure (PIT402) High High_Pre-Ignition" : Real = PLC "84_Setpoints".PIT402_Pilot_HighHigh AT %DB1.DBD0, 1 s
   "HMI Data_Inert Gas Pressure (PIT402) High_Post" : Real = PLC "84_Setpoints".PIT402_Post_High AT %DB1.DBD0, 1 s
   "HMI Data_Inert Gas Pressure (PIT402) High_Pre-Ignition" : Real = PLC "84_Setpoints".PIT402_Pilot_High AT %DB1.DBD0, 1 s
   "HMI Data_Inert Gas Pressure (PIT402) Low" : Real = PLC "84_Setpoints".PIT402_Main_Low AT %DB1.DBD0, 1 s
   "HMI Data_Inert Gas Pressure (PIT402) Low Low" : Real = PLC "84_Setpoints".PIT402_Main_LowLow AT %DB1.DBD0, 1 s
   "HMI Data_Inert Gas Pressure (PIT402) Low Low_Post" : Real = PLC "84_Setpoints".PIT402_Post_LowLow AT %DB1.DBD0, 1 s
   "HMI Data_Inert Gas Pressure (PIT402) Low Low_Pre-Ignition" : Real = PLC "84_Setpoints".PIT402_Pilot_LowLow AT %DB1.DBD0, 1 s
   "HMI Data_Inert Gas Pressure (PIT402) Low_Post" : Real = PLC "84_Setpoints".PIT402_Post_Low AT %DB1.DBD0, 1 s
   "HMI Data_Inert Gas Pressure (PIT402) Low_Pre-Ignition" : Real = PLC "84_Setpoints".PIT402_Pilot_Low AT %DB1.DBD0, 1 s
   "HMI Data_Inert Gas Temp (TIT401) High" : Real = PLC "84_Setpoints".TIT401_High AT %DB1.DBD0, 1 s
   "HMI Data_Inert Gas Temp (TIT401) High High" : Real = PLC "84_Setpoints".TIT401_HighHigh AT %DB1.DBD0, 1 s
   "HMI Data_Inlet CSW Pressure (PIT359) High" : Real = PLC "84_Setpoints".PIT359_High AT %DB1.DBD0, 1 s
   "HMI Data_Inlet CSW Pressure (PIT359) High High" : Real = PLC "84_Setpoints".PIT359_HighHigh AT %DB1.DBD0, 1 s
   "HMI Data_Inlet CSW Pressure (PIT359) Low" : Real = PLC "84_Setpoints".PIT359_Low AT %DB1.DBD0, 1 s
   "HMI Data_Inlet CSW Pressure (PIT359) Low Low" : Real = PLC "84_Setpoints".PIT359_LowLow AT %DB1.DBD0, 1 s
   "HMI Data_Inlet IA Pressure (PIT112) High" : Real = PLC "84_Setpoints".PIT112_High AT %DB1.DBD0, 1 s
   "HMI Data_Inlet IA Pressure (PIT112) High High" : Real = PLC "84_Setpoints".PIT112_HighHigh AT %DB1.DBD0, 1 s
   "HMI Data_Inlet IA Pressure (PIT112) Low" : Real = PLC "84_Setpoints".PIT112_Low AT %DB1.DBD0, 1 s
   "HMI Data_Inlet IA Pressure (PIT112) Low Low" : Real = PLC "84_Setpoints".PIT112_LowLow AT %DB1.DBD0, 1 s
   "HMI Data_Main Burner Fuel Pressure High" : Real = PLC "84_Setpoints".PIT205_High AT %DB1.DBD0, 1 s
   "HMI Data_Main Burner Fuel Pressure High High" : Real = PLC "84_Setpoints".PIT205_HighHigh AT %DB1.DBD0, 1 s
   "HMI Data_Main Burner Fuel Pressure Low" : Real = PLC "84_Setpoints".PIT205_Low AT %DB1.DBD0, 1 s
   "HMI Data_Main Burner Fuel Pressure Low Low SP" : Real = PLC "84_Setpoints".PIT205_LowLow AT %DB1.DBD0, 1 s
   "HMI Data_O2 Setpoint" : Real, internal
   "HMI Data_Outlet CSW Pressure (PIT316) High" : Real = PLC "84_Setpoints".PIT316_High AT %DB1.DBD0, 1 s
   "HMI Data_Outlet CSW Pressure (PIT316) High High" : Real = PLC "84_Setpoints".PIT316_HighHigh AT %DB1.DBD0, 1 s
   "HMI Data_Outlet CSW Pressure (PIT316) Low" : Real = PLC "84_Setpoints".PIT316_Low AT %DB1.DBD0, 1 s
   "HMI Data_Outlet CSW Pressure (PIT316) Low Low" : Real = PLC "84_Setpoints".PIT316_LowLow AT %DB1.DBD0, 1 s
   "HMI Data_PIT113 Target" : Real = PLC "84_Setpoints".PIT113_Pilot_Target AT %DB1.DBD0, 1 s
   "HMI Data_PIT205 Target" : Real = PLC "84_Setpoints".PIT205_Target AT %DB1.DBD0, 1 s
   "HMI Data_PIT402 Main Target" : Real = PLC "84_Setpoints".PIT402_Main_Target AT %DB1.DBD0, 1 s
   "HMI Data_PIT402 Pilot Target" : Real = PLC "84_Setpoints".PIT402_Pilot_Target AT %DB1.DBD0, 1 s
   "HMI Data_PIT402 Post Target Maximum" : Real = PLC "84_Setpoints".PIT401_Post_Target_Max AT %DB1.DBD0, 1 s
   "HMI Data_PIT402 Post Target Start" : Real = PLC "84_Setpoints".PIT402_Post_Target_Start AT %DB1.DBD0, 1 s
   "HMI Data_Shell CSW Temp High" : Real = PLC "84_Setpoints".TIT315_High AT %DB1.DBX0.0, 1 s
   "HMI Data_Shell CSW Temp High High" : Real = PLC "84_Setpoints".TIT315_HighHigh AT %DB1.DBD0, 1 s
   "HMI Data_Soot Content High" : Real = PLC "84_Setpoints".TX700_High AT %DB1.DBD0, 1 s
   "HMI Data_Soot Content Low" : Real = PLC "84_Setpoints".TX700_Low AT %DB1.DBD0, 1 s
   "HMI FAT Mode" : Bool = PLC "80_From_HMI".FAT_Mode AT %DB1.DBX0.0, 1 s
   "HMI Fuel Pump 1 Run Time" : LTime = PLC "82_To_HMI"."Run Time A" AT %DB1.DBD0, 1 s
   "HMI Fuel Pump 2 Run Time" : LTime = PLC "82_To_HMI"."Run Time B" AT %DB1.DBD0, 1 s
   "HMI Fuel Pump Duty Select" : Bool = PLC "80_From_HMI".SW_DTY_PMP_E500 AT %DB1.DBW0, 1 s
   "HMI Fuel Pump Service Reset" : Bool = PLC "80_From_HMI".RST_E500A_RT AT %DB1.DBX0.0, 1 s
   "HMI Indication Logic_DB_FA Mode Selected" : Bool = PLC "HMI Indication Logic_DB"."FA Mode Selected", 1 s
   "HMI Indication Logic_DB_Sequence Finished" : Bool = PLC "HMI Indication Logic_DB"."Sequence Finished", 1 s
   "HMI Indication Logic_DB_Tank Selected" : Bool = PLC "HMI Indication Logic_DB"."Tank Selected", 1 s
   "HMI Reset Auto" : Bool = PLC "80_From_HMI".RST_AUT_SEQ AT %DB1.DBX0.0, 1 s
   "HMI Standalone IGG" : Bool = PLC "80_From_HMI".IGG_STND_ALN AT %DB1.DBX0.0, 1 s
   "HMI Start IGGS" : Bool = PLC "80_From_HMI".RUN_IGG AT %DB1.DBX0.0, 1 s
   "HMI Stop IGGS" : Bool = PLC "80_From_HMI".STOP_IGG AT %DB1.DBX0.0, 1 s
   "I&A Compressor Run Hours" : Int = PLC "82_To_HMI"."I&A Compressor Run Hours", 1 s
   "I&A Compressor Run Minutes" : Int = PLC "82_To_HMI"."I&A Compressor Run Minutes", 1 s
   "I&A Compressor Run Seconds" : Int = PLC "82_To_HMI"."I&A Compressor Run Seconds", 1 s
   "I&A Compressor Total Run Hours" : Int = PLC "82_To_HMI"."I&A Compressor Run Hours", 1 s
   "IA Comp Control" : Bool = PLC "14_DQ_Data".E131ControlOut AT %DB1.DBX0.0, 1 s
   "IA Comp Warning" : Bool = PLC "10 DI_DATA".E131_WRNG AT %DB1.DBX0.0, 1 s
   "IA Compressor Animation" : Int = PLC "82_To_HMI"."IA Compressor Animation", 1 s
   "IA Compressor Healthy" : Bool = PLC "10 DI_DATA".E131_OK AT %DB1.DBX0.0, 1 s